   END_IF;
   IF #_w1 AND ("DB-PrioridadesCmpAlta".Vcmp3 = "DB-PrioridadesCmpAlta".Vcmp2) THEN
       "DB-PrioridadesCmpAlta".Vcmp2 := "DB-PrioridadesCmpAlta".Vcmp2 + 1;
   END_IF;
   IF #_w1 AND ("DB-PrioridadesCmpAlta".Vcmp3 = "DB-PrioridadesCmpAlta".Vcmp4) THEN
       "DB-PrioridadesCmpAlta".Vcmp4 := "DB-PrioridadesCmpAlta".Vcmp4 + 1;
   END_IF;
   IF #_w1 AND ("DB-PrioridadesCmpAlta".Vcmp3 = "DB-PrioridadesCmpAlta".Vcmp5) THEN
       "DB-PrioridadesCmpAlta".Vcmp5 := "DB-PrioridadesCmpAlta".Vcmp5 + 1;
   END_IF;
   IF #_w1 AND ("DB-PrioridadesCmpAlta".Vcmp3 = "DB-PrioridadesCmpAlta".Vcmp6) THEN
       "DB-PrioridadesCmpAlta".Vcmp6 := "DB-PrioridadesCmpAlta".Vcmp6 + 1;
   END_IF;
END_REGION

REGION Network 7
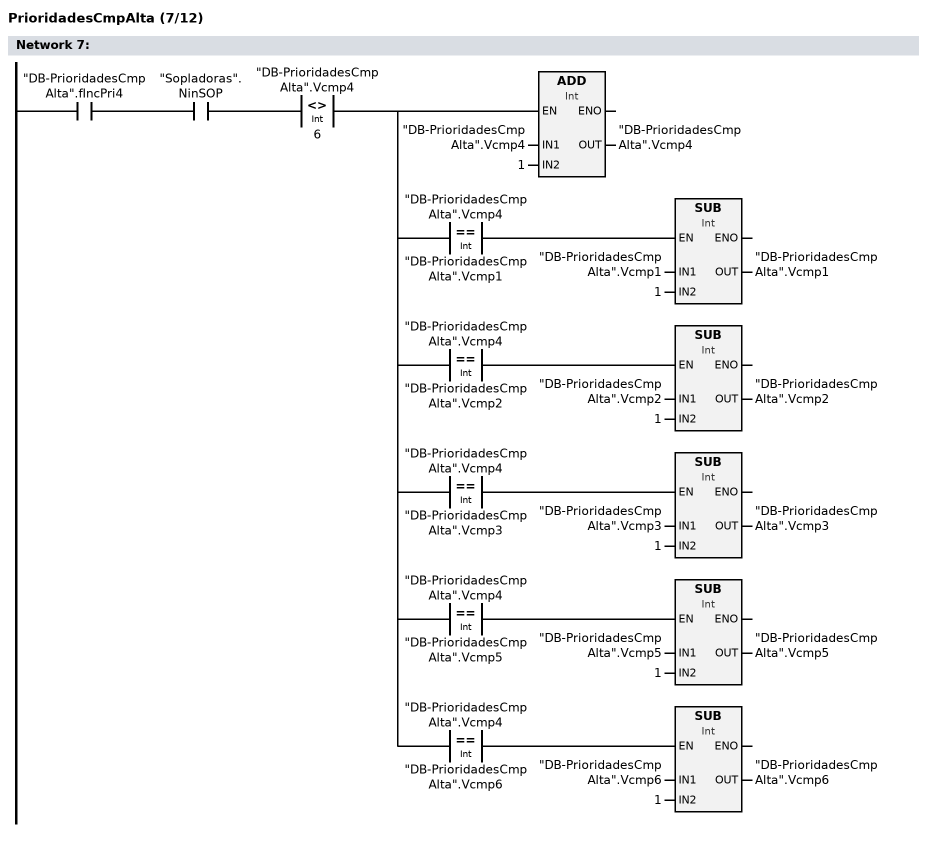
   RUNG wire#powerrail
      Contact( "DB-PrioridadesCmpAlta".fIncPri4 )
      Contact( "Sopladoras".NinSOP )
      { S7_Templates := "SrcType := Int" } NE_Contact(in1 := "DB-PrioridadesCmpAlta".Vcmp4, in2 := 6)
      wire#w1
      { S7_Templates := "SrcType := Int"; S7_GenerateENO := "TRUE" } Add(in1 := "DB-PrioridadesCmpAlta".Vcmp4, in2 := 1, out => "DB-PrioridadesCmpAlta".Vcmp4)
   END_RUNG
   RUNG wire#w1
      { S7_Templates := "SrcType := Int" } EQ_Contact(in1 := "DB-PrioridadesCmpAlta".Vcmp4, in2 := "DB-PrioridadesCmpAlta".Vcmp1)
      { S7_Templates := "SrcType := Int"; S7_GenerateENO := "TRUE" } Sub(in1 := "DB-PrioridadesCmpAlta".Vcmp1, in2 := 1, out => "DB-PrioridadesCmpAlta".Vcmp1)
   END_RUNG
   RUNG wire#w1
      { S7_Templates := "SrcType := Int" } EQ_Contact(in1 := "DB-PrioridadesCmpAlta".Vcmp4, in2 := "DB-PrioridadesCmpAlta".Vcmp2)
      { S7_Templates := "SrcType := Int"; S7_GenerateENO := "TRUE" } Sub(in1 := "DB-PrioridadesCmpAlta".Vcmp2, in2 := 1, out => "DB-PrioridadesCmpAlta".Vcmp2)
   END_RUNG
   RUNG wire#w1
      { S7_Templates := "SrcType := Int" } EQ_Contact(in1 := "DB-PrioridadesCmpAlta".Vcmp4, in2 := "DB-PrioridadesCmpAlta".Vcmp3)
      { S7_Templates := "SrcType := Int"; S7_GenerateENO := "TRUE" } Sub(in1 := "DB-PrioridadesCmpAlta".Vcmp3, in2 := 1, out => "DB-PrioridadesCmpAlta".Vcmp3)
   END_RUNG
   RUNG wire#w1
      { S7_Templates := "SrcType := Int" } EQ_Contact(in1 := "DB-PrioridadesCmpAlta".Vcmp4, in2 := "DB-PrioridadesCmpAlta".Vcmp5)
      { S7_Templates := "SrcType := Int"; S7_GenerateENO := "TRUE" } Sub(in1 := "DB-PrioridadesCmpAlta".Vcmp5, in2 := 1, out => "DB-PrioridadesCmpAlta".Vcmp5)
   END_RUNG
   RUNG wire#w1
      { S7_Templates := "SrcType := Int" } EQ_Contact(in1 := "DB-PrioridadesCmpAlta".Vcmp4, in2 := "DB-PrioridadesCmpAlta".Vcmp6)
      { S7_Templates := "SrcType := Int"; S7_GenerateENO := "TRUE" } Sub(in1 := "DB-PrioridadesCmpAlta".Vcmp6, in2 := 1, out => "DB-PrioridadesCmpAlta".Vcmp6)
   END_RUNG
   // the same network as SCL:
   #_w1 := "DB-PrioridadesCmpAlta".fIncPri4 AND "Sopladoras".NinSOP AND ("DB-PrioridadesCmpAlta".Vcmp4 <> 6);
   IF #_w1 THEN "DB-PrioridadesCmpAlta".Vcmp4 := "DB-PrioridadesCmpAlta".Vcmp4 + 1; END_IF;
   IF #_w1 AND ("DB-PrioridadesCmpAlta".Vcmp4 = "DB-PrioridadesCmpAlta".Vcmp1) THEN
       "DB-PrioridadesCmpAlta".Vcmp1 := "DB-PrioridadesCmpAlta".Vcmp1 - 1;
   END_IF;
   IF #_w1 AND ("DB-PrioridadesCmpAlta".Vcmp4 = "DB-PrioridadesCmpAlta".Vcmp2) THEN
       "DB-PrioridadesCmpAlta".Vcmp2 := "DB-PrioridadesCmpAlta".Vcmp2 - 1;
   END_IF;
   IF #_w1 AND ("DB-PrioridadesCmpAlta".Vcmp4 = "DB-PrioridadesCmpAlta".Vcmp3) THEN
       "DB-PrioridadesCmpAlta".Vcmp3 := "DB-PrioridadesCmpAlta".Vcmp3 - 1;
   END_IF;
   IF #_w1 AND ("DB-PrioridadesCmpAlta".Vcmp4 = "DB-PrioridadesCmpAlta".Vcmp5) THEN
       "DB-PrioridadesCmpAlta".Vcmp5 := "DB-PrioridadesCmpAlta".Vcmp5 - 1;
   END_IF;
   IF #_w1 AND ("DB-PrioridadesCmpAlta".Vcmp4 = "DB-PrioridadesCmpAlta".Vcmp6) THEN
       "DB-PrioridadesCmpAlta".Vcmp6 := "DB-PrioridadesCmpAlta".Vcmp6 - 1;
   END_IF;
END_REGION

REGION Network 8
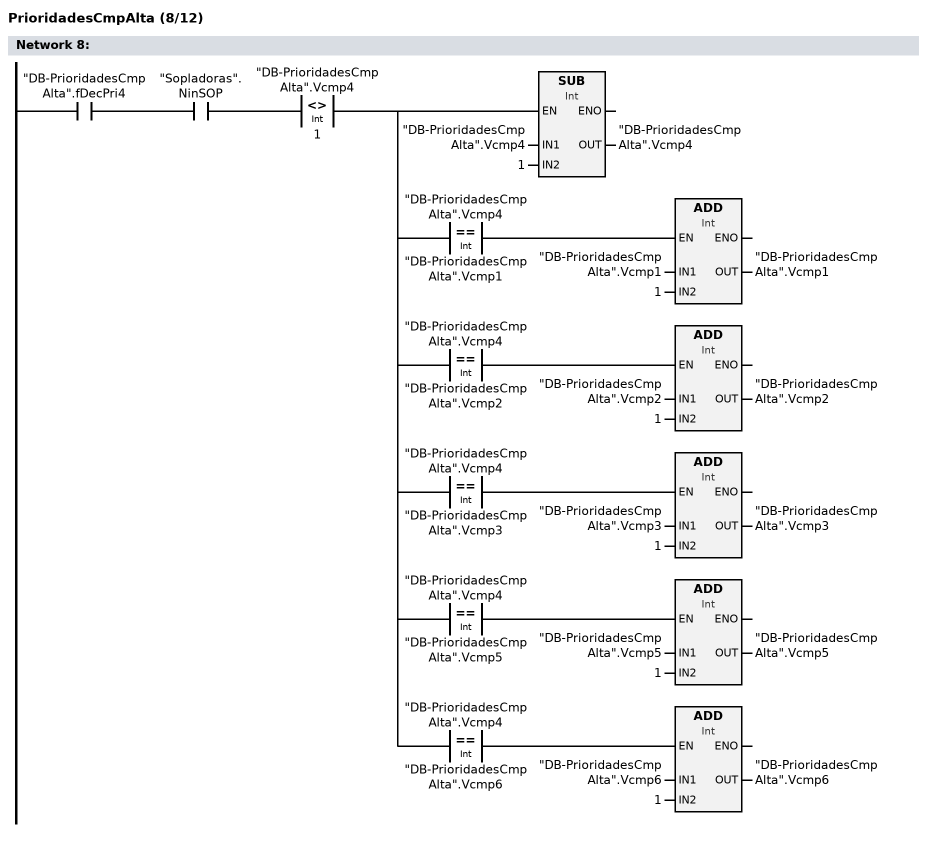
   RUNG wire#powerrail
      Contact( "DB-PrioridadesCmpAlta".fDecPri4 )
      Contact( "Sopladoras".NinSOP )
      { S7_Templates := "SrcType := Int" } NE_Contact(in1 := "DB-PrioridadesCmpAlta".Vcmp4, in2 := 1)
      wire#w1
      { S7_Templates := "SrcType := Int"; S7_GenerateENO := "TRUE" } Sub(in1 := "DB-PrioridadesCmpAlta".Vcmp4, in2 := 1, out => "DB-PrioridadesCmpAlta".Vcmp4)
   END_RUNG
   RUNG wire#w1
      { S7_Templates := "SrcType := Int" } EQ_Contact(in1 := "DB-PrioridadesCmpAlta".Vcmp4, in2 := "DB-PrioridadesCmpAlta".Vcmp1)
      { S7_Templates := "SrcType := Int"; S7_GenerateENO := "TRUE" } Add(in1 := "DB-PrioridadesCmpAlta".Vcmp1, in2 := 1, out => "DB-PrioridadesCmpAlta".Vcmp1)
   END_RUNG
   RUNG wire#w1
      { S7_Templates := "SrcType := Int" } EQ_Contact(in1 := "DB-PrioridadesCmpAlta".Vcmp4, in2 := "DB-PrioridadesCmpAlta".Vcmp2)
      { S7_Templates := "SrcType := Int"; S7_GenerateENO := "TRUE" } Add(in1 := "DB-PrioridadesCmpAlta".Vcmp2, in2 := 1, out => "DB-PrioridadesCmpAlta".Vcmp2)
   END_RUNG
   RUNG wire#w1
      { S7_Templates := "SrcType := Int" } EQ_Contact(in1 := "DB-PrioridadesCmpAlta".Vcmp4, in2 := "DB-PrioridadesCmpAlta".Vcmp3)
      { S7_Templates := "SrcType := Int"; S7_GenerateENO := "TRUE" } Add(in1 := "DB-PrioridadesCmpAlta".Vcmp3, in2 := 1, out => "DB-PrioridadesCmpAlta".Vcmp3)
   END_RUNG
   RUNG wire#w1
      { S7_Templates := "SrcType := Int" } EQ_Contact(in1 := "DB-PrioridadesCmpAlta".Vcmp4, in2 := "DB-PrioridadesCmpAlta".Vcmp5)
      { S7_Templates := "SrcType := Int"; S7_GenerateENO := "TRUE" } Add(in1 := "DB-PrioridadesCmpAlta".Vcmp5, in2 := 1, out => "DB-PrioridadesCmpAlta".Vcmp5)
   END_RUNG
   RUNG wire#w1
      { S7_Templates := "SrcType := Int" } EQ_Contact(in1 := "DB-PrioridadesCmpAlta".Vcmp4, in2 := "DB-PrioridadesCmpAlta".Vcmp6)
      { S7_Templates := "SrcType := Int"; S7_GenerateENO := "TRUE" } Add(in1 := "DB-PrioridadesCmpAlta".Vcmp6, in2 := 1, out => "DB-PrioridadesCmpAlta".Vcmp6)
   END_RUNG
   // the same network as SCL:
   #_w1 := "DB-PrioridadesCmpAlta".fDecPri4 AND "Sopladoras".NinSOP AND ("DB-PrioridadesCmpAlta".Vcmp4 <> 1);
   IF #_w1 THEN "DB-PrioridadesCmpAlta".Vcmp4 := "DB-PrioridadesCmpAlta".Vcmp4 - 1; END_IF;
   IF #_w1 AND ("DB-PrioridadesCmpAlta".Vcmp4 = "DB-PrioridadesCmpAlta".Vcmp1) THEN
       "DB-PrioridadesCmpAlta".Vcmp1 := "DB-PrioridadesCmpAlta".Vcmp1 + 1;
   END_IF;
   IF #_w1 AND ("DB-PrioridadesCmpAlta".Vcmp4 = "DB-PrioridadesCmpAlta".Vcmp2) THEN
       "DB-PrioridadesCmpAlta".Vcmp2 := "DB-PrioridadesCmpAlta".Vcmp2 + 1;
   END_IF;
   IF #_w1 AND ("DB-PrioridadesCmpAlta".Vcmp4 = "DB-PrioridadesCmpAlta".Vcmp3) THEN
       "DB-PrioridadesCmpAlta".Vcmp3 := "DB-PrioridadesCmpAlta".Vcmp3 + 1;
   END_IF;
   IF #_w1 AND ("DB-PrioridadesCmpAlta".Vcmp4 = "DB-PrioridadesCmpAlta".Vcmp5) THEN
       "DB-PrioridadesCmpAlta".Vcmp5 := "DB-PrioridadesCmpAlta".Vcmp5 + 1;
   END_IF;
   IF #_w1 AND ("DB-PrioridadesCmpAlta".Vcmp4 = "DB-PrioridadesCmpAlta".Vcmp6) THEN
       "DB-PrioridadesCmpAlta".Vcmp6 := "DB-PrioridadesCmpAlta".Vcmp6 + 1;
   END_IF;
END_REGION

REGION Network 9
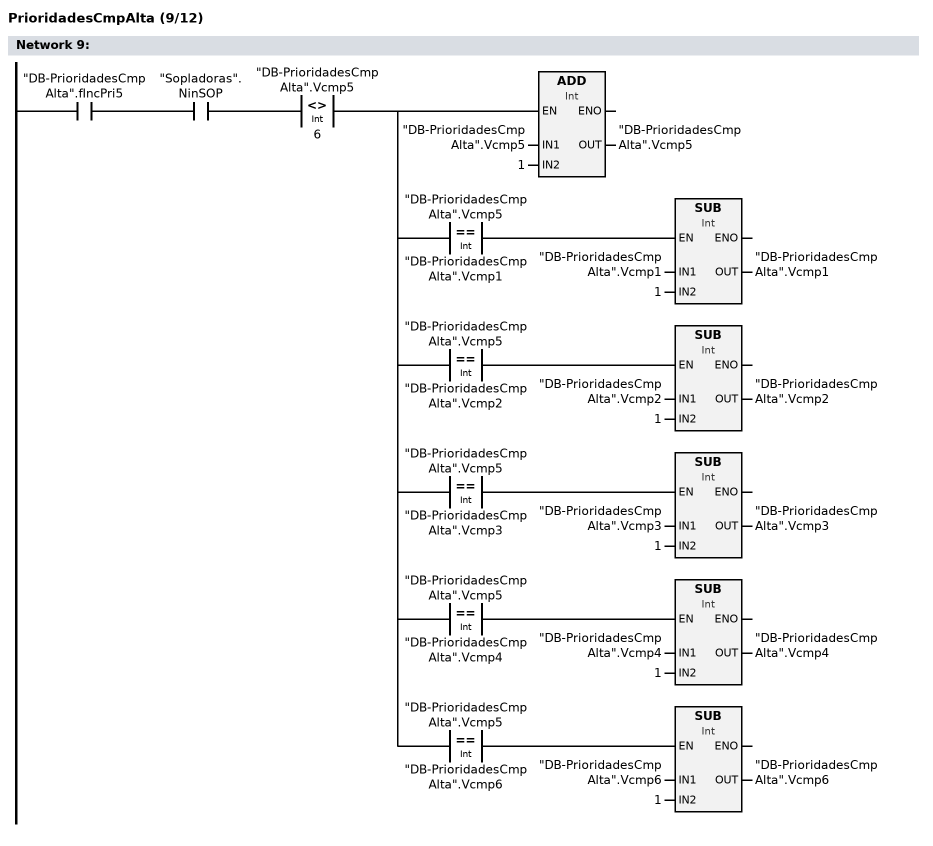
   RUNG wire#powerrail
      Contact( "DB-PrioridadesCmpAlta".fIncPri5 )
      Contact( "Sopladoras".NinSOP )
      { S7_Templates := "SrcType := Int" } NE_Contact(in1 := "DB-PrioridadesCmpAlta".Vcmp5, in2 := 6)
      wire#w1
      { S7_Templates := "SrcType := Int"; S7_GenerateENO := "TRUE" } Add(in1 := "DB-PrioridadesCmpAlta".Vcmp5, in2 := 1, out => "DB-PrioridadesCmpAlta".Vcmp5)
   END_RUNG
   RUNG wire#w1
      { S7_Templates := "SrcType := Int" } EQ_Contact(in1 := "DB-PrioridadesCmpAlta".Vcmp5, in2 := "DB-PrioridadesCmpAlta".Vcmp1)
      { S7_Templates := "SrcType := Int"; S7_GenerateENO := "TRUE" } Sub(in1 := "DB-PrioridadesCmpAlta".Vcmp1, in2 := 1, out => "DB-PrioridadesCmpAlta".Vcmp1)
   END_RUNG
   RUNG wire#w1
      { S7_Templates := "SrcType := Int" } EQ_Contact(in1 := "DB-PrioridadesCmpAlta".Vcmp5, in2 := "DB-PrioridadesCmpAlta".Vcmp2)
      { S7_Templates := "SrcType := Int"; S7_GenerateENO := "TRUE" } Sub(in1 := "DB-PrioridadesCmpAlta".Vcmp2, in2 := 1, out => "DB-PrioridadesCmpAlta".Vcmp2)
   END_RUNG
   RUNG wire#w1
      { S7_Templates := "SrcType := Int" } EQ_Contact(in1 := "DB-PrioridadesCmpAlta".Vcmp5, in2 := "DB-PrioridadesCmpAlta".Vcmp3)
      { S7_Templates := "SrcType := Int"; S7_GenerateENO := "TRUE" } Sub(in1 := "DB-PrioridadesCmpAlta".Vcmp3, in2 := 1, out => "DB-PrioridadesCmpAlta".Vcmp3)
   END_RUNG
   RUNG wire#w1
      { S7_Templates := "SrcType := Int" } EQ_Contact(in1 := "DB-PrioridadesCmpAlta".Vcmp5, in2 := "DB-PrioridadesCmpAlta".Vcmp4)
      { S7_Templates := "SrcType := Int"; S7_GenerateENO := "TRUE" } Sub(in1 := "DB-PrioridadesCmpAlta".Vcmp4, in2 := 1, out => "DB-PrioridadesCmpAlta".Vcmp4)
   END_RUNG
   RUNG wire#w1
      { S7_Templates := "SrcType := Int" } EQ_Contact(in1 := "DB-PrioridadesCmpAlta".Vcmp5, in2 := "DB-PrioridadesCmpAlta".Vcmp6)
      { S7_Templates := "SrcType := Int"; S7_GenerateENO := "TRUE" } Sub(in1 := "DB-PrioridadesCmpAlta".Vcmp6, in2 := 1, out => "DB-PrioridadesCmpAlta".Vcmp6)
   END_RUNG
   // the same network as SCL:
   #_w1 := "DB-PrioridadesCmpAlta".fIncPri5 AND "Sopladoras".NinSOP AND ("DB-PrioridadesCmpAlta".Vcmp5 <> 6);
   IF #_w1 THEN "DB-PrioridadesCmpAlta".Vcmp5 := "DB-PrioridadesCmpAlta".Vcmp5 + 1; END_IF;
   IF #_w1 AND ("DB-PrioridadesCmpAlta".Vcmp5 = "DB-PrioridadesCmpAlta".Vcmp1) THEN
       "DB-PrioridadesCmpAlta".Vcmp1 := "DB-PrioridadesCmpAlta".Vcmp1 - 1;
   END_IF;
   IF #_w1 AND ("DB-PrioridadesCmpAlta".Vcmp5 = "DB-PrioridadesCmpAlta".Vcmp2) THEN
       "DB-PrioridadesCmpAlta".Vcmp2 := "DB-PrioridadesCmpAlta".Vcmp2 - 1;
   END_IF;
   IF #_w1 AND ("DB-PrioridadesCmpAlta".Vcmp5 = "DB-PrioridadesCmpAlta".Vcmp3) THEN
       "DB-PrioridadesCmpAlta".Vcmp3 := "DB-PrioridadesCmpAlta".Vcmp3 - 1;
   END_IF;
   IF #_w1 AND ("DB-PrioridadesCmpAlta".Vcmp5 = "DB-PrioridadesCmpAlta".Vcmp4) THEN
       "DB-PrioridadesCmpAlta".Vcmp4 := "DB-PrioridadesCmpAlta".Vcmp4 - 1;
   END_IF;
   IF #_w1 AND ("DB-PrioridadesCmpAlta".Vcmp5 = "DB-PrioridadesCmpAlta".Vcmp6) THEN
       "DB-PrioridadesCmpAlta".Vcmp6 := "DB-PrioridadesCmpAlta".Vcmp6 - 1;
   END_IF;
END_REGION

REGION Network 10
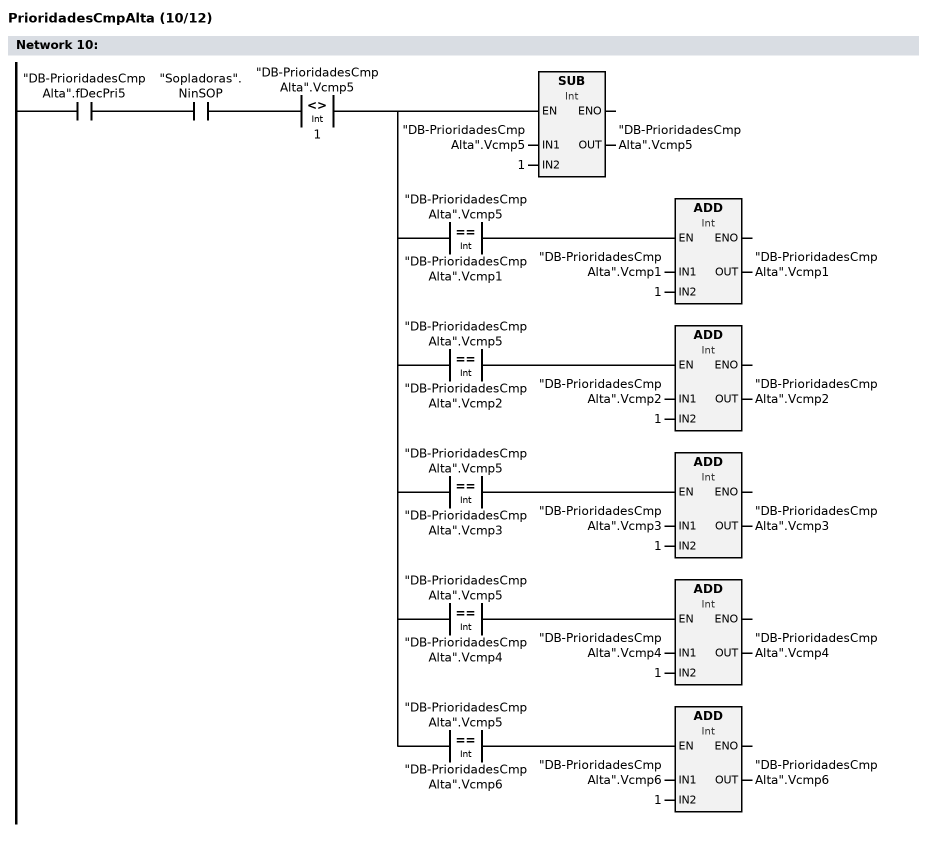
   RUNG wire#powerrail
      Contact( "DB-PrioridadesCmpAlta".fDecPri5 )
      Contact( "Sopladoras".NinSOP )
      { S7_Templates := "SrcType := Int" } NE_Contact(in1 := "DB-PrioridadesCmpAlta".Vcmp5, in2 := 1)
      wire#w1
      { S7_Templates := "SrcType := Int"; S7_GenerateENO := "TRUE" } Sub(in1 := "DB-PrioridadesCmpAlta".Vcmp5, in2 := 1, out => "DB-PrioridadesCmpAlta".Vcmp5)
   END_RUNG
   RUNG wire#w1
      { S7_Templates := "SrcType := Int" } EQ_Contact(in1 := "DB-PrioridadesCmpAlta".Vcmp5, in2 := "DB-PrioridadesCmpAlta".Vcmp1)
      { S7_Templates := "SrcType := Int"; S7_GenerateENO := "TRUE" } Add(in1 := "DB-PrioridadesCmpAlta".Vcmp1, in2 := 1, out => "DB-PrioridadesCmpAlta".Vcmp1)
   END_RUNG
   RUNG wire#w1
      { S7_Templates := "SrcType := Int" } EQ_Contact(in1 := "DB-PrioridadesCmpAlta".Vcmp5, in2 := "DB-PrioridadesCmpAlta".Vcmp2)
      { S7_Templates := "SrcType := Int"; S7_GenerateENO := "TRUE" } Add(in1 := "DB-PrioridadesCmpAlta".Vcmp2, in2 := 1, out => "DB-PrioridadesCmpAlta".Vcmp2)
   END_RUNG
   RUNG wire#w1
      { S7_Templates := "SrcType := Int" } EQ_Contact(in1 := "DB-PrioridadesCmpAlta".Vcmp5, in2 := "DB-PrioridadesCmpAlta".Vcmp3)
      { S7_Templates := "SrcType := Int"; S7_GenerateENO := "TRUE" } Add(in1 := "DB-PrioridadesCmpAlta".Vcmp3, in2 := 1, out => "DB-PrioridadesCmpAlta".Vcmp3)
   END_RUNG
   RUNG wire#w1
      { S7_Templates := "SrcType := Int" } EQ_Contact(in1 := "DB-PrioridadesCmpAlta".Vcmp5, in2 := "DB-PrioridadesCmpAlta".Vcmp4)
      { S7_Templates := "SrcType := Int"; S7_GenerateENO := "TRUE" } Add(in1 := "DB-PrioridadesCmpAlta".Vcmp4, in2 := 1, out => "DB-PrioridadesCmpAlta".Vcmp4)
   END_RUNG
   RUNG wire#w1
      { S7_Templates := "SrcType := Int" } EQ_Contact(in1 := "DB-PrioridadesCmpAlta".Vcmp5, in2 := "DB-PrioridadesCmpAlta".Vcmp6)
      { S7_Templates := "SrcType := Int"; S7_GenerateENO := "TRUE" } Add(in1 := "DB-PrioridadesCmpAlta".Vcmp6, in2 := 1, out => "DB-PrioridadesCmpAlta".Vcmp6)
   END_RUNG
   // the same network as SCL:
   #_w1 := "DB-PrioridadesCmpAlta".fDecPri5 AND "Sopladoras".NinSOP AND ("DB-PrioridadesCmpAlta".Vcmp5 <> 1);
   IF #_w1 THEN "DB-PrioridadesCmpAlta".Vcmp5 := "DB-PrioridadesCmpAlta".Vcmp5 - 1; END_IF;
   IF #_w1 AND ("DB-PrioridadesCmpAlta".Vcmp5 = "DB-PrioridadesCmpAlta".Vcmp1) THEN
       "DB-PrioridadesCmpAlta".Vcmp1 := "DB-PrioridadesCmpAlta".Vcmp1 + 1;
   END_IF;
   IF #_w1 AND ("DB-PrioridadesCmpAlta".Vcmp5 = "DB-PrioridadesCmpAlta".Vcmp2) THEN
       "DB-PrioridadesCmpAlta".Vcmp2 := "DB-PrioridadesCmpAlta".Vcmp2 + 1;
   END_IF;
   IF #_w1 AND ("DB-PrioridadesCmpAlta".Vcmp5 = "DB-PrioridadesCmpAlta".Vcmp3) THEN
       "DB-PrioridadesCmpAlta".Vcmp3 := "DB-PrioridadesCmpAlta".Vcmp3 + 1;
   END_IF;
   IF #_w1 AND ("DB-PrioridadesCmpAlta".Vcmp5 = "DB-PrioridadesCmpAlta".Vcmp4) THEN
       "DB-PrioridadesCmpAlta".Vcmp4 := "DB-PrioridadesCmpAlta".Vcmp4 + 1;
   END_IF;
   IF #_w1 AND ("DB-PrioridadesCmpAlta".Vcmp5 = "DB-PrioridadesCmpAlta".Vcmp6) THEN
       "DB-PrioridadesCmpAlta".Vcmp6 := "DB-PrioridadesCmpAlta".Vcmp6 + 1;
   END_IF;
END_REGION

REGION Network 11
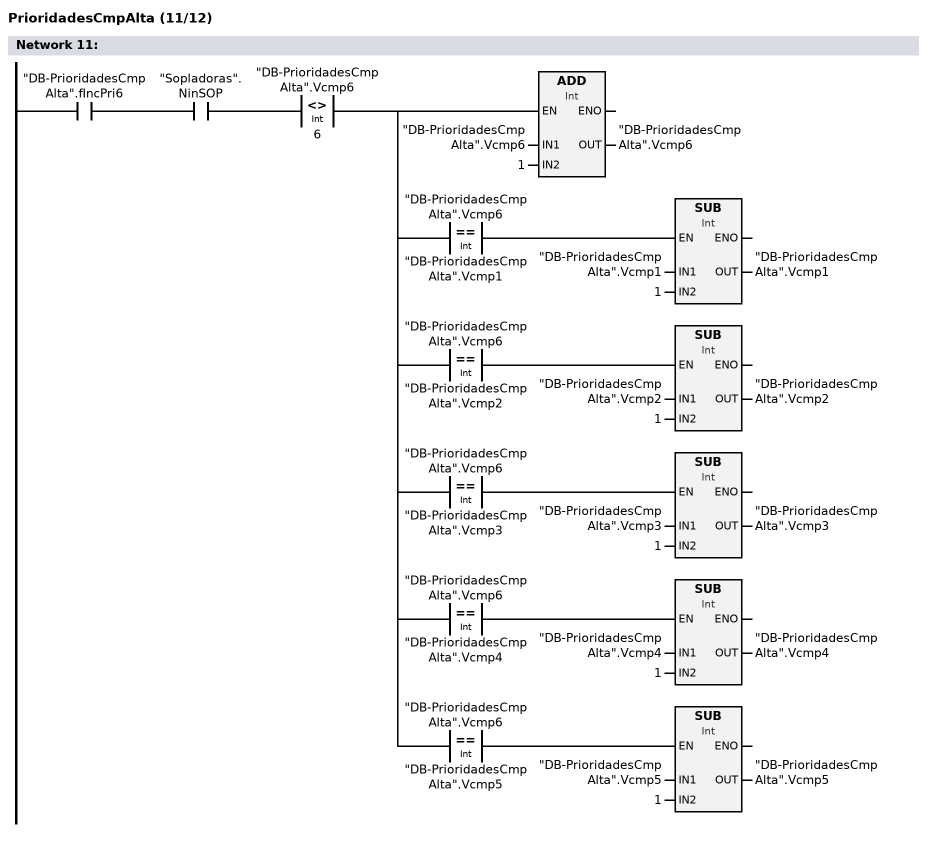
   RUNG wire#powerrail
      Contact( "DB-PrioridadesCmpAlta".fIncPri6 )
      Contact( "Sopladoras".NinSOP )
      { S7_Templates := "SrcType := Int" } NE_Contact(in1 := "DB-PrioridadesCmpAlta".Vcmp6, in2 := 6)
      wire#w1
      { S7_Templates := "SrcType := Int"; S7_GenerateENO := "TRUE" } Add(in1 := "DB-PrioridadesCmpAlta".Vcmp6, in2 := 1, out => "DB-PrioridadesCmpAlta".Vcmp6)
   END_RUNG
   RUNG wire#w1
      { S7_Templates := "SrcType := Int" } EQ_Contact(in1 := "DB-PrioridadesCmpAlta".Vcmp6, in2 := "DB-PrioridadesCmpAlta".Vcmp1)
      { S7_Templates := "SrcType := Int"; S7_GenerateENO := "TRUE" } Sub(in1 := "DB-PrioridadesCmpAlta".Vcmp1, in2 := 1, out => "DB-PrioridadesCmpAlta".Vcmp1)
   END_RUNG
   RUNG wire#w1
      { S7_Templates := "SrcType := Int" } EQ_Contact(in1 := "DB-PrioridadesCmpAlta".Vcmp6, in2 := "DB-PrioridadesCmpAlta".Vcmp2)
      { S7_Templates := "SrcType := Int"; S7_GenerateENO := "TRUE" } Sub(in1 := "DB-PrioridadesCmpAlta".Vcmp2, in2 := 1, out => "DB-PrioridadesCmpAlta".Vcmp2)
   END_RUNG
   RUNG wire#w1
      { S7_Templates := "SrcType := Int" } EQ_Contact(in1 := "DB-PrioridadesCmpAlta".Vcmp6, in2 := "DB-PrioridadesCmpAlta".Vcmp3)
      { S7_Templates := "SrcType := Int"; S7_GenerateENO := "TRUE" } Sub(in1 := "DB-PrioridadesCmpAlta".Vcmp3, in2 := 1, out => "DB-PrioridadesCmpAlta".Vcmp3)
   END_RUNG
   RUNG wire#w1
      { S7_Templates := "SrcType := Int" } EQ_Contact(in1 := "DB-PrioridadesCmpAlta".Vcmp6, in2 := "DB-PrioridadesCmpAlta".Vcmp4)
      { S7_Templates := "SrcType := Int"; S7_GenerateENO := "TRUE" } Sub(in1 := "DB-PrioridadesCmpAlta".Vcmp4, in2 := 1, out => "DB-PrioridadesCmpAlta".Vcmp4)
   END_RUNG
   RUNG wire#w1
      { S7_Templates := "SrcType := Int" } EQ_Contact(in1 := "DB-PrioridadesCmpAlta".Vcmp6, in2 := "DB-PrioridadesCmpAlta".Vcmp5)
      { S7_Templates := "SrcType := Int"; S7_GenerateENO := "TRUE" } Sub(in1 := "DB-PrioridadesCmpAlta".Vcmp5, in2 := 1, out => "DB-PrioridadesCmpAlta".Vcmp5)
   END_RUNG
   // the same network as SCL:
   #_w1 := "DB-PrioridadesCmpAlta".fIncPri6 AND "Sopladoras".NinSOP AND ("DB-PrioridadesCmpAlta".Vcmp6 <> 6);
   IF #_w1 THEN "DB-PrioridadesCmpAlta".Vcmp6 := "DB-PrioridadesCmpAlta".Vcmp6 + 1; END_IF;
   IF #_w1 AND ("DB-PrioridadesCmpAlta".Vcmp6 = "DB-PrioridadesCmpAlta".Vcmp1) THEN
       "DB-PrioridadesCmpAlta".Vcmp1 := "DB-PrioridadesCmpAlta".Vcmp1 - 1;
   END_IF;
   IF #_w1 AND ("DB-PrioridadesCmpAlta".Vcmp6 = "DB-PrioridadesCmpAlta".Vcmp2) THEN
       "DB-PrioridadesCmpAlta".Vcmp2 := "DB-PrioridadesCmpAlta".Vcmp2 - 1;
   END_IF;
   IF #_w1 AND ("DB-PrioridadesCmpAlta".Vcmp6 = "DB-PrioridadesCmpAlta".Vcmp3) THEN
       "DB-PrioridadesCmpAlta".Vcmp3 := "DB-PrioridadesCmpAlta".Vcmp3 - 1;
   END_IF;
   IF #_w1 AND ("DB-PrioridadesCmpAlta".Vcmp6 = "DB-PrioridadesCmpAlta".Vcmp4) THEN
       "DB-PrioridadesCmpAlta".Vcmp4 := "DB-PrioridadesCmpAlta".Vcmp4 - 1;
   END_IF;
   IF #_w1 AND ("DB-PrioridadesCmpAlta".Vcmp6 = "DB-PrioridadesCmpAlta".Vcmp5) THEN
       "DB-PrioridadesCmpAlta".Vcmp5 := "DB-PrioridadesCmpAlta".Vcmp5 - 1;
   END_IF;
END_REGION

REGION Network 12
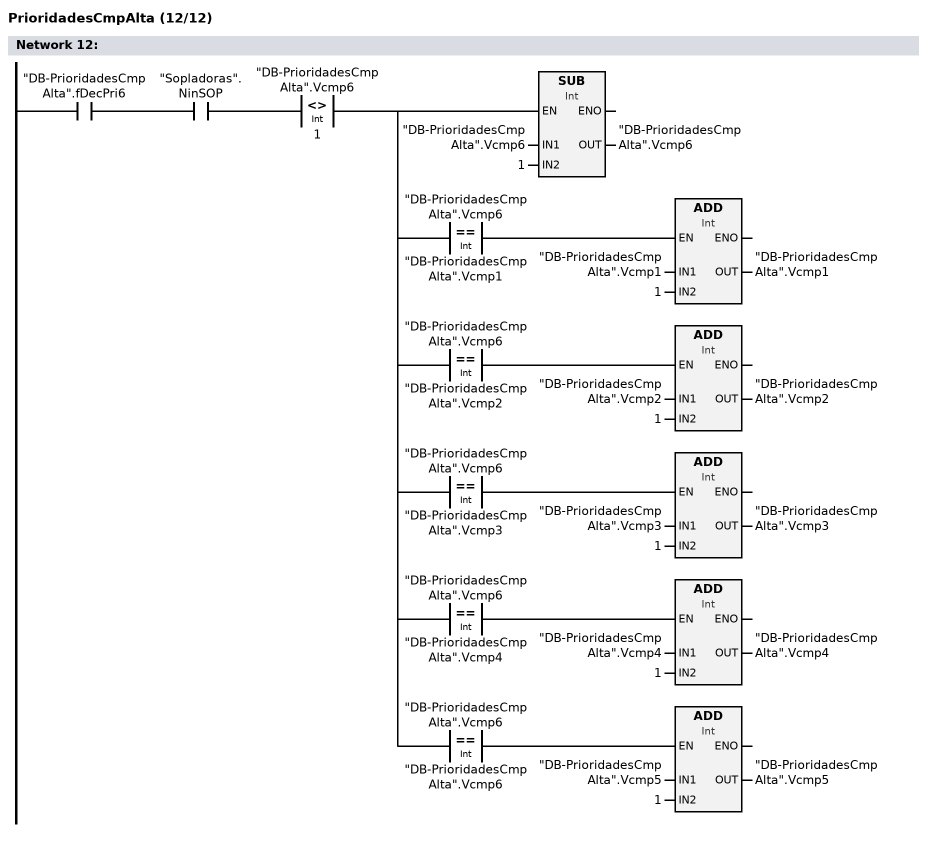
   RUNG wire#powerrail
      Contact( "DB-PrioridadesCmpAlta".fDecPri6 )
      Contact( "Sopladoras".NinSOP )
      { S7_Templates := "SrcType := Int" } NE_Contact(in1 := "DB-PrioridadesCmpAlta".Vcmp6, in2 := 1)
      wire#w1
      { S7_Templates := "SrcType := Int"; S7_GenerateENO := "TRUE" } Sub(in1 := "DB-PrioridadesCmpAlta".Vcmp6, in2 := 1, out => "DB-PrioridadesCmpAlta".Vcmp6)
   END_RUNG
   RUNG wire#w1
      { S7_Templates := "SrcType := Int" } EQ_Contact(in1 := "DB-PrioridadesCmpAlta".Vcmp6, in2 := "DB-PrioridadesCmpAlta".Vcmp1)
      { S7_Templates := "SrcType := Int"; S7_GenerateENO := "TRUE" } Add(in1 := "DB-PrioridadesCmpAlta".Vcmp1, in2 := 1, out => "DB-PrioridadesCmpAlta".Vcmp1)
   END_RUNG
   RUNG wire#w1
      { S7_Templates := "SrcType := Int" } EQ_Contact(in1 := "DB-PrioridadesCmpAlta".Vcmp6, in2 := "DB-PrioridadesCmpAlta".Vcmp2)
      { S7_Templates := "SrcType := Int"; S7_GenerateENO := "TRUE" } Add(in1 := "DB-PrioridadesCmpAlta".Vcmp2, in2 := 1, out => "DB-PrioridadesCmpAlta".Vcmp2)
   END_RUNG
   RUNG wire#w1
      { S7_Templates := "SrcType := Int" } EQ_Contact(in1 := "DB-PrioridadesCmpAlta".Vcmp6, in2 := "DB-PrioridadesCmpAlta".Vcmp3)
      { S7_Templates := "SrcType := Int"; S7_GenerateENO := "TRUE" } Add(in1 := "DB-PrioridadesCmpAlta".Vcmp3, in2 := 1, out => "DB-PrioridadesCmpAlta".Vcmp3)
   END_RUNG
   RUNG wire#w1
      { S7_Templates := "SrcType := Int" } EQ_Contact(in1 := "DB-PrioridadesCmpAlta".Vcmp6, in2 := "DB-PrioridadesCmpAlta".Vcmp4)
      { S7_Templates := "SrcType := Int"; S7_GenerateENO := "TRUE" } Add(in1 := "DB-PrioridadesCmpAlta".Vcmp4, in2 := 1, out => "DB-PrioridadesCmpAlta".Vcmp4)
   END_RUNG
   RUNG wire#w1
      { S7_Templates := "SrcType := Int" } EQ_Contact(in1 := "DB-PrioridadesCmpAlta".Vcmp6, in2 := "DB-PrioridadesCmpAlta".Vcmp6)
      { S7_Templates := "SrcType := Int"; S7_GenerateENO := "TRUE" } Add(in1 := "DB-PrioridadesCmpAlta".Vcmp5, in2 := 1, out => "DB-PrioridadesCmpAlta".Vcmp5)
   END_RUNG
   // the same network as SCL:
   #_w1 := "DB-PrioridadesCmpAlta".fDecPri6 AND "Sopladoras".NinSOP AND ("DB-PrioridadesCmpAlta".Vcmp6 <> 1);
   IF #_w1 THEN "DB-PrioridadesCmpAlta".Vcmp6 := "DB-PrioridadesCmpAlta".Vcmp6 - 1; END_IF;
   IF #_w1 AND ("DB-PrioridadesCmpAlta".Vcmp6 = "DB-PrioridadesCmpAlta".Vcmp1) THEN
       "DB-PrioridadesCmpAlta".Vcmp1 := "DB-PrioridadesCmpAlta".Vcmp1 + 1;
   END_IF;
   IF #_w1 AND ("DB-PrioridadesCmpAlta".Vcmp6 = "DB-PrioridadesCmpAlta".Vcmp2) THEN
       "DB-PrioridadesCmpAlta".Vcmp2 := "DB-PrioridadesCmpAlta".Vcmp2 + 1;
   END_IF;
   IF #_w1 AND ("DB-PrioridadesCmpAlta".Vcmp6 = "DB-PrioridadesCmpAlta".Vcmp3) THEN
       "DB-PrioridadesCmpAlta".Vcmp3 := "DB-PrioridadesCmpAlta".Vcmp3 + 1;
   END_IF;
   IF #_w1 AND ("DB-PrioridadesCmpAlta".Vcmp6 = "DB-PrioridadesCmpAlta".Vcmp4) THEN
       "DB-PrioridadesCmpAlta".Vcmp4 := "DB-PrioridadesCmpAlta".Vcmp4 + 1;
   END_IF;
   IF #_w1 AND ("DB-PrioridadesCmpAlta".Vcmp6 = "DB-PrioridadesCmpAlta".Vcmp6) THEN
       "DB-PrioridadesCmpAlta".Vcmp5 := "DB-PrioridadesCmpAlta".Vcmp5 + 1;
   END_IF;
END_REGION
END_FUNCTION

FUNCTION "AccionamientosCmpAlta" : Void   // FC34, LAD
{ S7_Optimized_Access := 'FALSE' }
VERSION : 0.1
   VAR_TEMP   // added for the SCL form of the ladder/FBD networks
      _w1 : Bool;
      _s5time1 : S5Time;
   END_VAR
BEGIN

REGION Network 1: Dejar abrir valvula compresor 1 / Habilitación para poner en carga compresor de alta ABC2
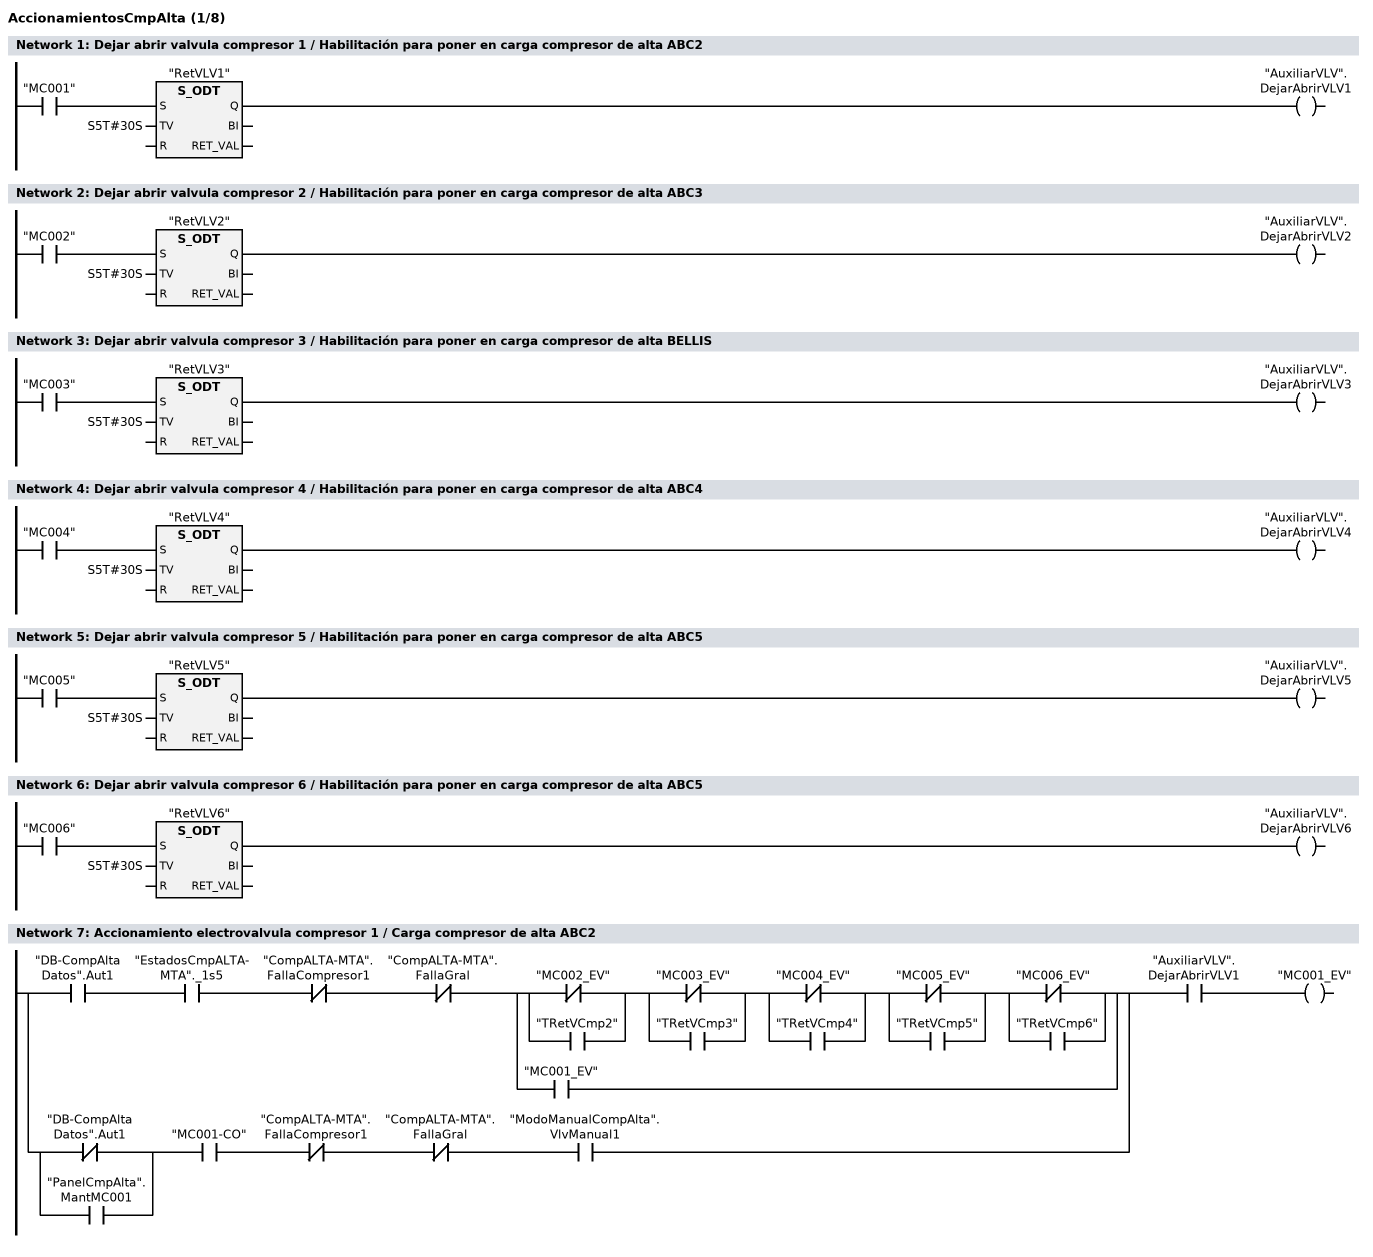
   RUNG wire#powerrail
      Contact( "MC001" )
      S_ODT(T_NO := "RetVLV1", TV := S5T#30S, R :=, BI =>, RET_VAL =>)
      Coil( "AuxiliarVLV".DejarAbrirVLV1 )
   END_RUNG
   // the same network as SCL:
   #_s5time1 := S_ODT(T_NO := "RetVLV1", S := "MC001", TV := S5T#30S, Q => #_w1);
   "AuxiliarVLV".DejarAbrirVLV1 := #_w1;
END_REGION

REGION Network 2: Dejar abrir valvula compresor 2 / Habilitación para poner en carga compresor de alta ABC3
   RUNG wire#powerrail
      Contact( "MC002" )
      S_ODT(T_NO := "RetVLV2", TV := S5T#30S, R :=, BI =>, RET_VAL =>)
      Coil( "AuxiliarVLV".DejarAbrirVLV2 )
   END_RUNG
   // the same network as SCL:
   #_s5time1 := S_ODT(T_NO := "RetVLV2", S := "MC002", TV := S5T#30S, Q => #_w1);
   "AuxiliarVLV".DejarAbrirVLV2 := #_w1;
END_REGION

REGION Network 3: Dejar abrir valvula compresor 3 / Habilitación para poner en carga compresor de alta BELLIS
   RUNG wire#powerrail
      Contact( "MC003" )
      S_ODT(T_NO := "RetVLV3", TV := S5T#30S, R :=, BI =>, RET_VAL =>)
      Coil( "AuxiliarVLV".DejarAbrirVLV3 )
   END_RUNG
   // the same network as SCL:
   #_s5time1 := S_ODT(T_NO := "RetVLV3", S := "MC003", TV := S5T#30S, Q => #_w1);
   "AuxiliarVLV".DejarAbrirVLV3 := #_w1;
END_REGION

REGION Network 4: Dejar abrir valvula compresor 4 / Habilitación para poner en carga compresor de alta ABC4
   RUNG wire#powerrail
      Contact( "MC004" )
      S_ODT(T_NO := "RetVLV4", TV := S5T#30S, R :=, BI =>, RET_VAL =>)
      Coil( "AuxiliarVLV".DejarAbrirVLV4 )
   END_RUNG
   // the same network as SCL:
   #_s5time1 := S_ODT(T_NO := "RetVLV4", S := "MC004", TV := S5T#30S, Q => #_w1);
   "AuxiliarVLV".DejarAbrirVLV4 := #_w1;
END_REGION

REGION Network 5: Dejar abrir valvula compresor 5 / Habilitación para poner en carga compresor de alta ABC5
   RUNG wire#powerrail
      Contact( "MC005" )
      S_ODT(T_NO := "RetVLV5", TV := S5T#30S, R :=, BI =>, RET_VAL =>)
      Coil( "AuxiliarVLV".DejarAbrirVLV5 )
   END_RUNG
   // the same network as SCL:
   #_s5time1 := S_ODT(T_NO := "RetVLV5", S := "MC005", TV := S5T#30S, Q => #_w1);
   "AuxiliarVLV".DejarAbrirVLV5 := #_w1;
END_REGION

REGION Network 6: Dejar abrir valvula compresor 6 / Habilitación para poner en carga compresor de alta ABC5
   RUNG wire#powerrail
      Contact( "MC006" )
      S_ODT(T_NO := "RetVLV6", TV := S5T#30S, R :=, BI =>, RET_VAL =>)
      Coil( "AuxiliarVLV".DejarAbrirVLV6 )
   END_RUNG
   // the same network as SCL:
   #_s5time1 := S_ODT(T_NO := "RetVLV6", S := "MC006", TV := S5T#30S, Q => #_w1);
   "AuxiliarVLV".DejarAbrirVLV6 := #_w1;
END_REGION

REGION Network 7: Accionamiento electrovalvula compresor 1 / Carga compresor de alta ABC2
   RUNG wire#powerrail
      Contact( "DB-CompAltaDatos".Aut1 )
      Contact( "EstadosCmpALTA-MTA"._1s5 )
      I_Contact( "CompALTA-MTA".FallaCompresor1 )
      I_Contact( "CompALTA-MTA".FallaGral )
      wire#w1
      I_Contact( "MC002_EV" )
      wire#w2
      I_Contact( "MC003_EV" )
      wire#w3
      I_Contact( "MC004_EV" )
      wire#w4
      I_Contact( "MC005_EV" )
      wire#w5
      I_Contact( "MC006_EV" )
      wire#w6
      Contact( "AuxiliarVLV".DejarAbrirVLV1 )
      Coil( "MC001_EV" )
   END_RUNG
   RUNG wire#w1
      Contact( "TRetVCmp2" )
   END_RUNG wire#w2
   RUNG wire#w2
      Contact( "TRetVCmp3" )
   END_RUNG wire#w3
   RUNG wire#w3
      Contact( "TRetVCmp4" )
   END_RUNG wire#w4
   RUNG wire#w4
      Contact( "TRetVCmp5" )
   END_RUNG wire#w5
   RUNG wire#w5
      Contact( "TRetVCmp6" )
   END_RUNG wire#w6
   RUNG wire#w1
      Contact( "MC001_EV" )
   END_RUNG wire#w6
   RUNG wire#powerrail
      I_Contact( "DB-CompAltaDatos".Aut1 )
      wire#w7
      Contact( "MC001-CO" )
      I_Contact( "CompALTA-MTA".FallaCompresor1 )
      I_Contact( "CompALTA-MTA".FallaGral )
      Contact( "ModoManualCompAlta".VlvManual1 )
   END_RUNG wire#w6
   RUNG wire#powerrail
      Contact( "PanelCmpAlta".MantMC001 )
   END_RUNG wire#w7
   // the same network as SCL:
   "MC001_EV" := (("DB-CompAltaDatos".Aut1 AND "EstadosCmpALTA-MTA"._1s5 AND NOT "CompALTA-MTA".FallaCompresor1 AND NOT "CompALTA-MTA".FallaGral AND (((NOT "MC002_EV" OR "TRetVCmp2") AND (NOT "MC003_EV" OR "TRetVCmp3") AND (NOT "MC004_EV" OR "TRetVCmp4") AND (NOT "MC005_EV" OR "TRetVCmp5") AND (NOT "MC006_EV" OR "TRetVCmp6")) OR "MC001_EV")) OR ((NOT "DB-CompAltaDatos".Aut1 OR "PanelCmpAlta".MantMC001) AND "MC001-CO" AND NOT "CompALTA-MTA".FallaCompresor1 AND NOT "CompALTA-MTA".FallaGral AND "ModoManualCompAlta".VlvManual1)) AND "AuxiliarVLV".DejarAbrirVLV1;
END_REGION

REGION Network 8: Accionamiento electrovalvula compresor 2 / Carga compresor de alta ABC3
